(* Logix 5000 project; controller NWGG 1756-L72 rev 35.12; software revision 35.00 *) (continued)

ADD_ON_INSTRUCTION AndcoAnalog   (* revision 1.0 *)
VAR_IN_OUT
   Andco_Values : udt_Andco_Values; {required}
   Andco_Motor_Open : BOOL; {required}
   Anco_Motor_Close : BOOL; {required}
END_VAR
VAR_INPUT
   AnalogValue : DINT; {access Read Only, required}
END_VAR
VAR
   tmr_Web_Watchdog : TIMER := (PRE := 30000); {access None}
   Cal_Open_Gate : BOOL; {access None}
   Cal_Close_Gate : BOOL; {access None}
   Motor_Wind_Down : DINT; {access None}
   Cal_Mid_Point : DINT; {access None}
   Cal_Preact : BOOL; {access None}
   Cal_Finish_Close_Gate : BOOL; {access None}
   tmr_Motor_Wind_Down : TIMER[8] := ([1].PRE := 1000, [2].PRE := 1000); {access None}
   New_Position : DINT; {access None}
   Move_Open : BOOL; {access None}
   Move_Close : BOOL; {access None}
   Adjusted_New_Position : DINT; {access None}
   Cal_Init_Bin_Closed : BOOL; {access None}
   tmrCalCloseGate : TIMER := (PRE := 55000); {access None}
   CurrentPosition : DINT; {access None}
   tmrCalOpenGate : TIMER := (PRE := 55000); {access None}
   CalReturnToPosition : BOOL; {access None}
   CalibratingGate : BOOL; {access None}
   onsStartCal : BOOL; {access None}
   sbCalGateClosed : BOOL; {access None}
   obCalGateClosed : BOOL; {access None}
   sbStartCal : BOOL; {access None}
   obStartCal : BOOL; {access None}
   sbCalGateOpened : BOOL; {access None}
   obCalGateOpened : BOOL; {access None}
END_VAR

ROUTINE Logic   (* ladder *)
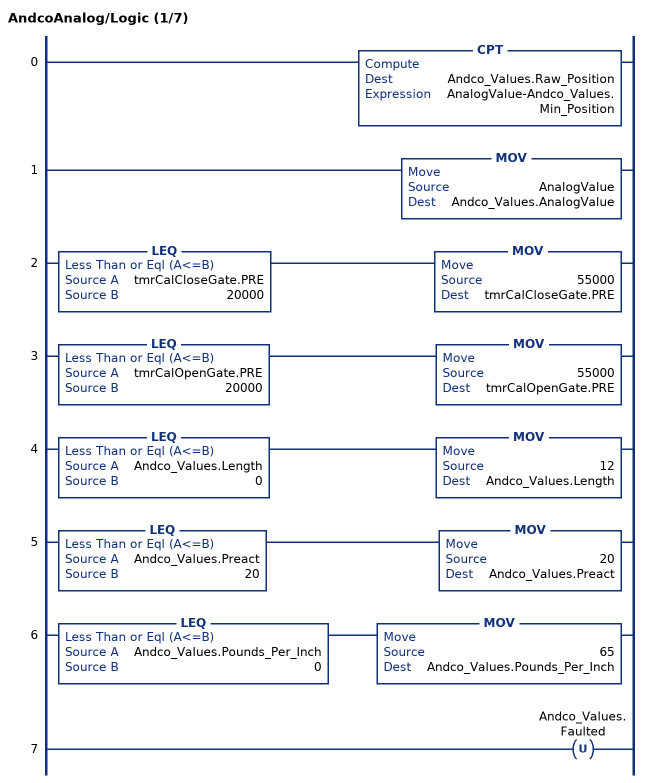
   0: CPT(Andco_Values.Raw_Position,AnalogValue-Andco_Values.Min_Position);
   1: MOV(AnalogValue,Andco_Values.AnalogValue);
   2: LEQ(tmrCalCloseGate.PRE,20000)MOV(55000,tmrCalCloseGate.PRE);
   3: LEQ(tmrCalOpenGate.PRE,20000)MOV(55000,tmrCalOpenGate.PRE);
   4: LEQ(Andco_Values.Length,0)MOV(12,Andco_Values.Length);
   5: LEQ(Andco_Values.Preact,20)MOV(20,Andco_Values.Preact);
   6: LEQ(Andco_Values.Pounds_Per_Inch,0)MOV(65,Andco_Values.Pounds_Per_Inch);
   7: OTU(Andco_Values.Faulted);
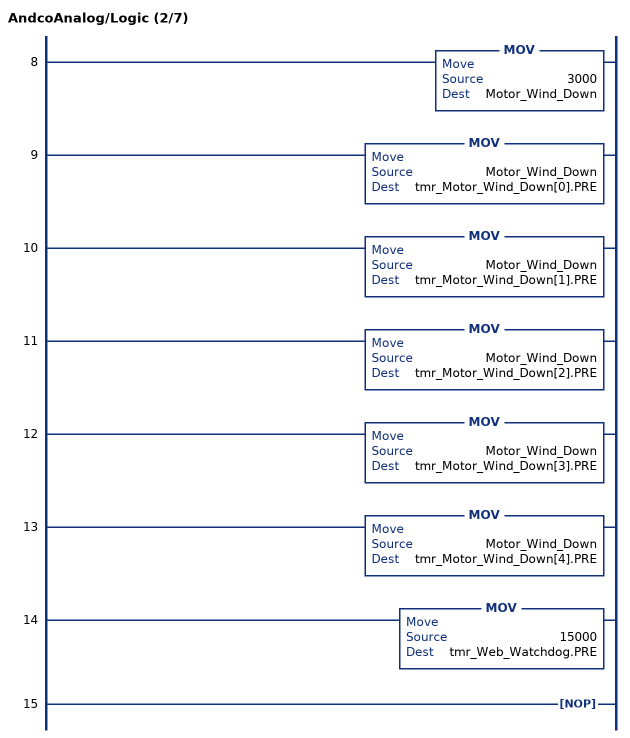
   8: MOV(3000,Motor_Wind_Down);
   9: MOV(Motor_Wind_Down,tmr_Motor_Wind_Down[0].PRE);
   10: MOV(Motor_Wind_Down,tmr_Motor_Wind_Down[1].PRE);
   11: MOV(Motor_Wind_Down,tmr_Motor_Wind_Down[2].PRE);
   12: MOV(Motor_Wind_Down,tmr_Motor_Wind_Down[3].PRE);
   13: MOV(Motor_Wind_Down,tmr_Motor_Wind_Down[4].PRE);
   14: MOV(15000,tmr_Web_Watchdog.PRE);
   15: NOP();
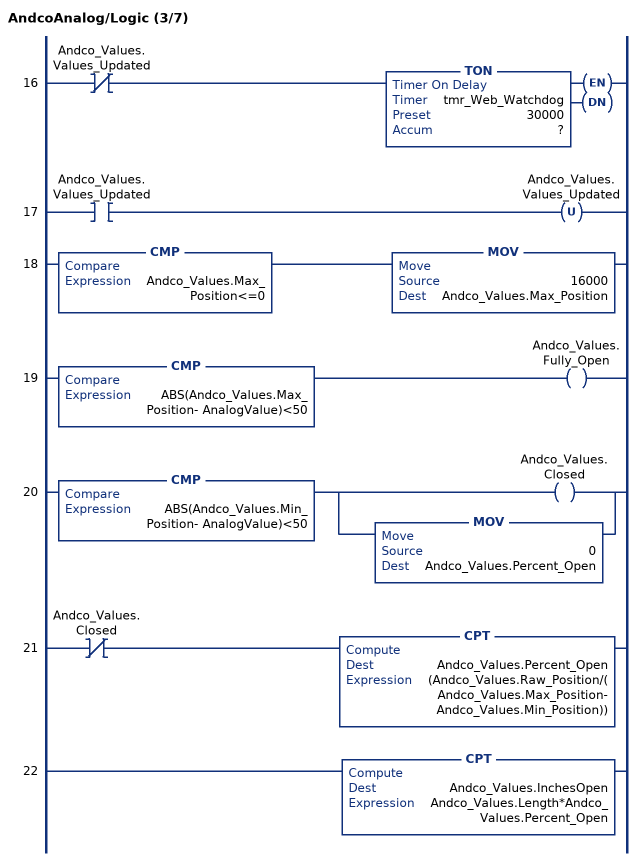
   16: XIO(Andco_Values.Values_Updated)TON(tmr_Web_Watchdog,?,?);
   17: XIC(Andco_Values.Values_Updated)OTU(Andco_Values.Values_Updated);
   18: CMP(Andco_Values.Max_Position<=0)MOV(16000,Andco_Values.Max_Position);
   19: CMP(ABS(Andco_Values.Max_Position- AnalogValue)<50)OTE(Andco_Values.Fully_Open);
   20: CMP(ABS(Andco_Values.Min_Position- AnalogValue)<50)[OTE(Andco_Values.Closed) ,MOV(0,Andco_Values.Percent_Open) ];
   21: XIO(Andco_Values.Closed)CPT(Andco_Values.Percent_Open,(Andco_Values.Raw_Position/(Andco_Values.Max_Position-Andco_Values.Min_Position)));
   22: CPT(Andco_Values.InchesOpen,Andco_Values.Length*Andco_Values.Percent_Open);
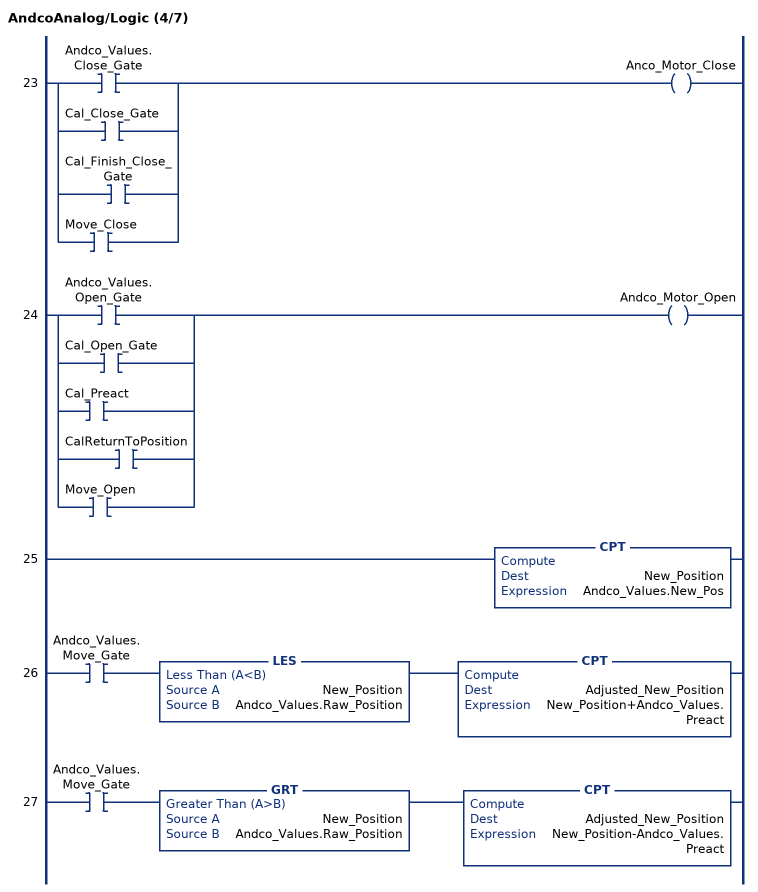
   23: [XIC(Andco_Values.Close_Gate) ,XIC(Cal_Close_Gate) ,XIC(Cal_Finish_Close_Gate) ,XIC(Move_Close) ]OTE(Anco_Motor_Close);
   24: [XIC(Andco_Values.Open_Gate) ,XIC(Cal_Open_Gate) ,XIC(Cal_Preact) ,XIC(CalReturnToPosition) ,XIC(Move_Open) ]OTE(Andco_Motor_Open);
   25: CPT(New_Position,Andco_Values.New_Pos);
   26: XIC(Andco_Values.Move_Gate)LES(New_Position,Andco_Values.Raw_Position)CPT(Adjusted_New_Position,New_Position+Andco_Values.Preact);
   27: XIC(Andco_Values.Move_Gate)GRT(New_Position,Andco_Values.Raw_Position)CPT(Adjusted_New_Position,New_Position-Andco_Values.Preact);
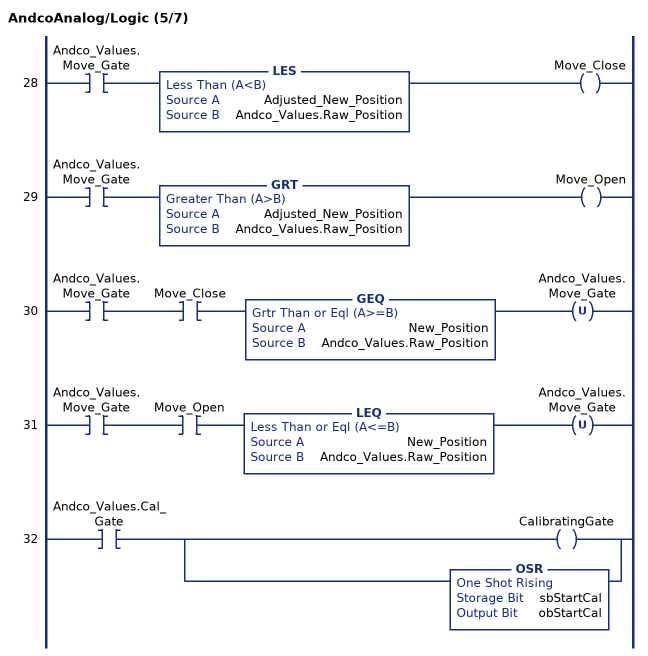
   28: XIC(Andco_Values.Move_Gate)LES(Adjusted_New_Position,Andco_Values.Raw_Position)OTE(Move_Close);
   29: XIC(Andco_Values.Move_Gate)GRT(Adjusted_New_Position,Andco_Values.Raw_Position)OTE(Move_Open);
   30: XIC(Andco_Values.Move_Gate)XIC(Move_Close)GEQ(New_Position,Andco_Values.Raw_Position)OTU(Andco_Values.Move_Gate);
   31: XIC(Andco_Values.Move_Gate)XIC(Move_Open)LEQ(New_Position,Andco_Values.Raw_Position)OTU(Andco_Values.Move_Gate);
   32: XIC(Andco_Values.Cal_Gate)[OTE(CalibratingGate) ,OSR(sbStartCal,obStartCal) ];
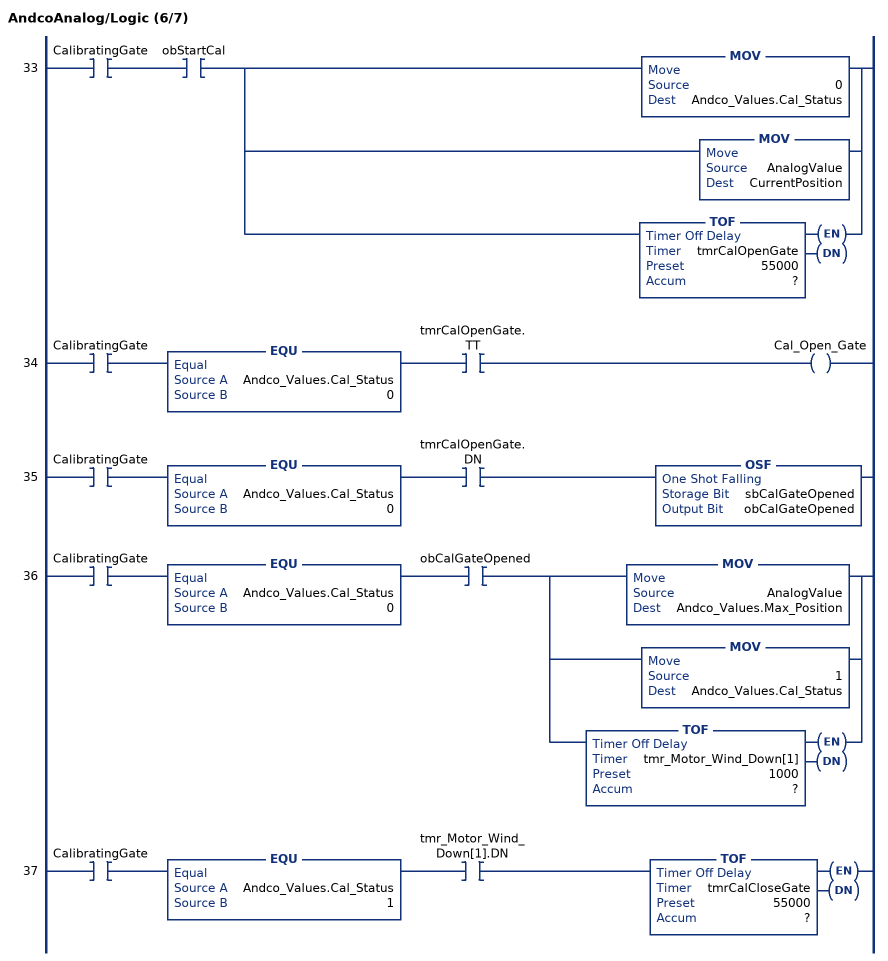
   33: XIC(CalibratingGate)XIC(obStartCal)[MOV(0,Andco_Values.Cal_Status) ,MOV(AnalogValue,CurrentPosition) ,TOF(tmrCalOpenGate,?,?) ];
   34: XIC(CalibratingGate)EQU(Andco_Values.Cal_Status,0)XIC(tmrCalOpenGate.TT)OTE(Cal_Open_Gate);
   35: XIC(CalibratingGate)EQU(Andco_Values.Cal_Status,0)XIC(tmrCalOpenGate.DN)OSF(sbCalGateOpened,obCalGateOpened);
   36: XIC(CalibratingGate)EQU(Andco_Values.Cal_Status,0)XIC(obCalGateOpened)[MOV(AnalogValue,Andco_Values.Max_Position) ,MOV(1,Andco_Values.Cal_Status) ,TOF(tmr_Motor_Wind_Down[1],?,?) ];
   37: XIC(CalibratingGate)EQU(Andco_Values.Cal_Status,1)XIC(tmr_Motor_Wind_Down[1].DN)TOF(tmrCalCloseGate,?,?);
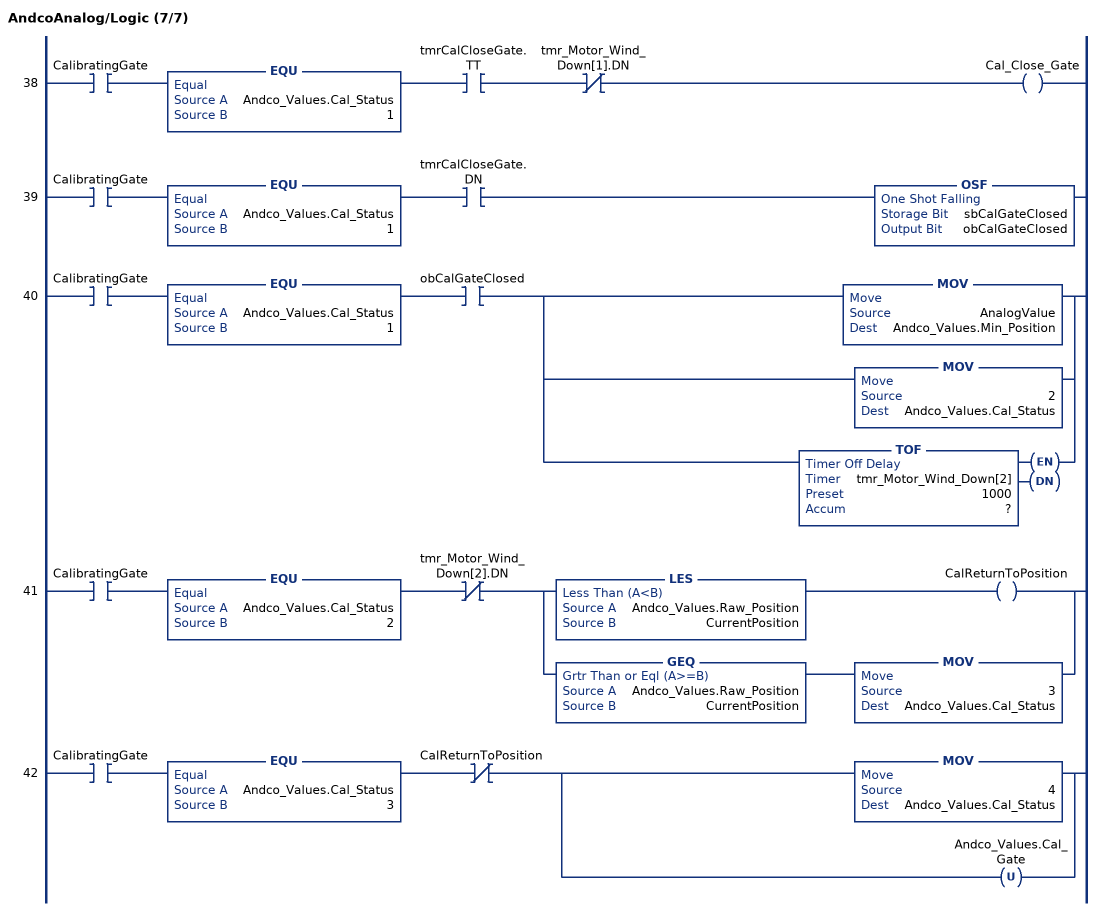
   38: XIC(CalibratingGate)EQU(Andco_Values.Cal_Status,1)XIC(tmrCalCloseGate.TT)XIO(tmr_Motor_Wind_Down[1].DN)OTE(Cal_Close_Gate);
   39: XIC(CalibratingGate)EQU(Andco_Values.Cal_Status,1)XIC(tmrCalCloseGate.DN)OSF(sbCalGateClosed,obCalGateClosed);
   40: XIC(CalibratingGate)EQU(Andco_Values.Cal_Status,1)XIC(obCalGateClosed)[MOV(AnalogValue,Andco_Values.Min_Position) ,MOV(2,Andco_Values.Cal_Status) ,TOF(tmr_Motor_Wind_Down[2],?,?) ];
   41: XIC(CalibratingGate)EQU(Andco_Values.Cal_Status,2)XIO(tmr_Motor_Wind_Down[2].DN)[LES(Andco_Values.Raw_Position,CurrentPosition) OTE(CalReturnToPosition) ,GEQ(Andco_Values.Raw_Position,CurrentPosition) MOV(3,Andco_Values.Cal_Status) ];
   42: XIC(CalibratingGate)EQU(Andco_Values.Cal_Status,3)XIO(CalReturnToPosition)[MOV(4,Andco_Values.Cal_Status) ,OTU(Andco_Values.Cal_Gate) ];
END_ROUTINE
END_ADD_ON_INSTRUCTION

ADD_ON_INSTRUCTION HOUR_METER   (* revision 1.0 *)
VAR_INPUT
   MOTOR_RUNNING_INPUT_1 : BOOL; {required}
END_VAR
VAR_OUTPUT
   HR_METER_DISPLAY : DINT; {visible}
END_VAR
VAR_INPUT
   NEXT_SCHDL_MAINTENANCE : DINT; {visible}
END_VAR
VAR_OUTPUT
   MAINTENANCE_ALARM : BOOL; {visible}
END_VAR
VAR
   COUNTER : COUNTER := (PRE := 99999999); {access None}
   TIMER : TIMER := (PRE := 3600000); {access None}
END_VAR

ROUTINE Logic   (* ladder *)
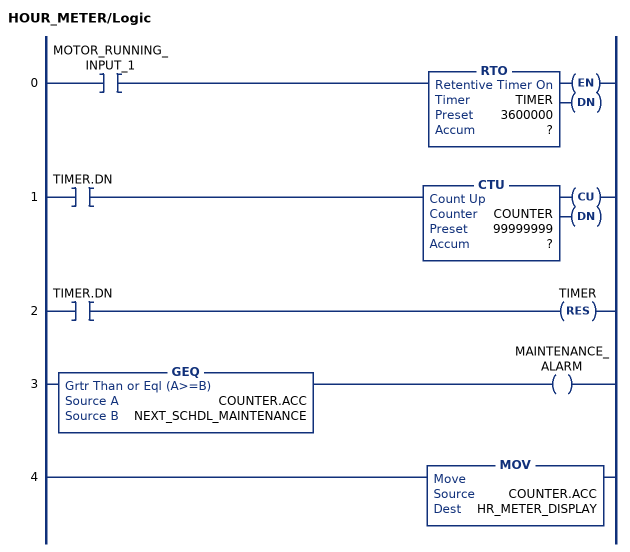
   0: XIC(MOTOR_RUNNING_INPUT_1)RTO(TIMER,?,?);
   1: XIC(TIMER.DN)CTU(COUNTER,?,?);
   2: XIC(TIMER.DN)RES(TIMER);
   3: GEQ(COUNTER.ACC,NEXT_SCHDL_MAINTENANCE)OTE(MAINTENANCE_ALARM);
   4: MOV(COUNTER.ACC,HR_METER_DISPLAY);
END_ROUTINE
END_ADD_ON_INSTRUCTION

ADD_ON_INSTRUCTION Loadout_Bin_Control   (* revision 1.0 *)
VAR_IN_OUT
   Bin : udt_Loadout_Bin; {required}
   Open_Air_Gate : BOOL; {required}
END_VAR
VAR_INPUT
   Bin_Open_Treat_Pause : BOOL; {required}
   Bin_Open_Clean_Pause : BOOL; {required}
END_VAR
VAR_IN_OUT
   TMR_Max_Treat_Delay : TIMER; {required}
   TMR_Max_Clean_Delay : TIMER; {required}
   Air_Gate_Open_Input : BOOL; {required}
   Auger_Relay : BOOL; {required}
END_VAR
VAR_INPUT
   Use_Auger_Relay : BOOL; {required}
   Use_Bindicator : BOOL; {access None, required}
END_VAR
VAR_IN_OUT
   Bindicator_Input : BOOL; {required}
   ALM_Air_Gate_Failed : ALARM_DIGITAL; {required}
END_VAR
VAR_INPUT
   Bin_Open_Transfer_Pause : BOOL; {required}
END_VAR
VAR_IN_OUT
   Clean_Batch_Status : DINT; {required}
   Treat_Batch_Status : DINT; {required}
   Transfer_Batch_Status : DINT; {required}
   Andco_Motor_Open : BOOL; {required}
   Andco_Motor_Close : BOOL; {required}
   Required_Belt : BOOL; {required}
   Manual_Mode : BOOL; {required}
END_VAR
VAR_INPUT
   RawAnalogTag : DINT; {access Read Only, required}
END_VAR
VAR
   Auto_Open_Air_Gate_Ready : BOOL; {access None}
   Air_Gate_Open_Cal : BOOL; {access None}
   TMR_Air_Gate_Fail : TIMER := (PRE := 4000); {access None}
   ALM_Air_Gate_Failed_Ack : BOOL; {access None}
   Air_Gate_Open_Clean : BOOL; {access None}
   Air_Gate_Open_Treat : BOOL; {access None}
   Air_Gate_Open_Transfer : BOOL; {access None}
   Andco : Andco; {access None}
   Open_Treat_Air_Gate : BOOL; {access None}
   Open_Treat_Air_Gate_Ready : BOOL; {access None}
   AndcoAnalog : AndcoAnalog; {access None}
END_VAR

ROUTINE Logic   (* ladder *)
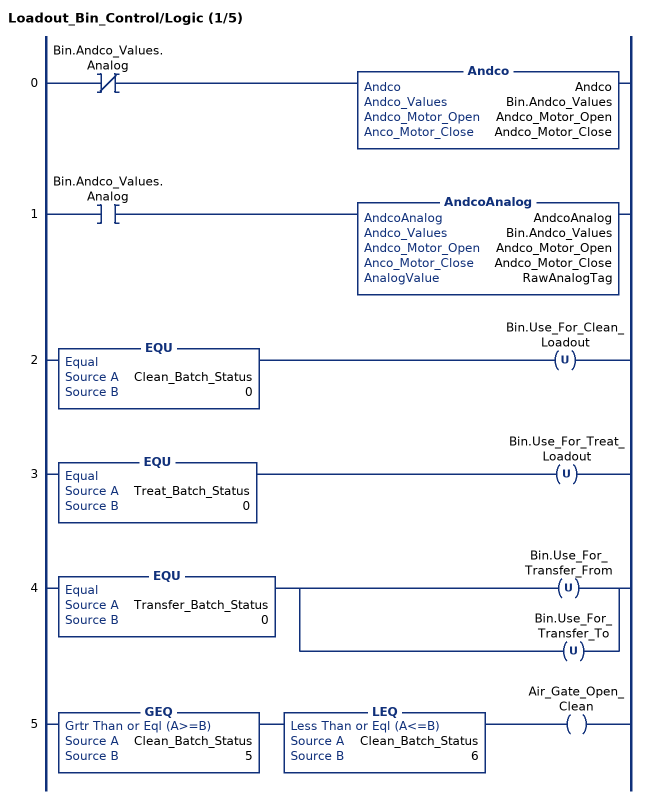
   0: XIO(Bin.Andco_Values.Analog)Andco(Andco,Bin.Andco_Values,Andco_Motor_Open,Andco_Motor_Close);
   1: XIC(Bin.Andco_Values.Analog)AndcoAnalog(AndcoAnalog,Bin.Andco_Values,Andco_Motor_Open,Andco_Motor_Close,RawAnalogTag);
   2: EQU(Clean_Batch_Status,0)OTU(Bin.Use_For_Clean_Loadout);
   3: EQU(Treat_Batch_Status,0)OTU(Bin.Use_For_Treat_Loadout);
   4: EQU(Transfer_Batch_Status,0)[OTU(Bin.Use_For_Transfer_From) ,OTU(Bin.Use_For_Transfer_To) ];
   5: GEQ(Clean_Batch_Status,5)LEQ(Clean_Batch_Status,6)OTE(Air_Gate_Open_Clean);
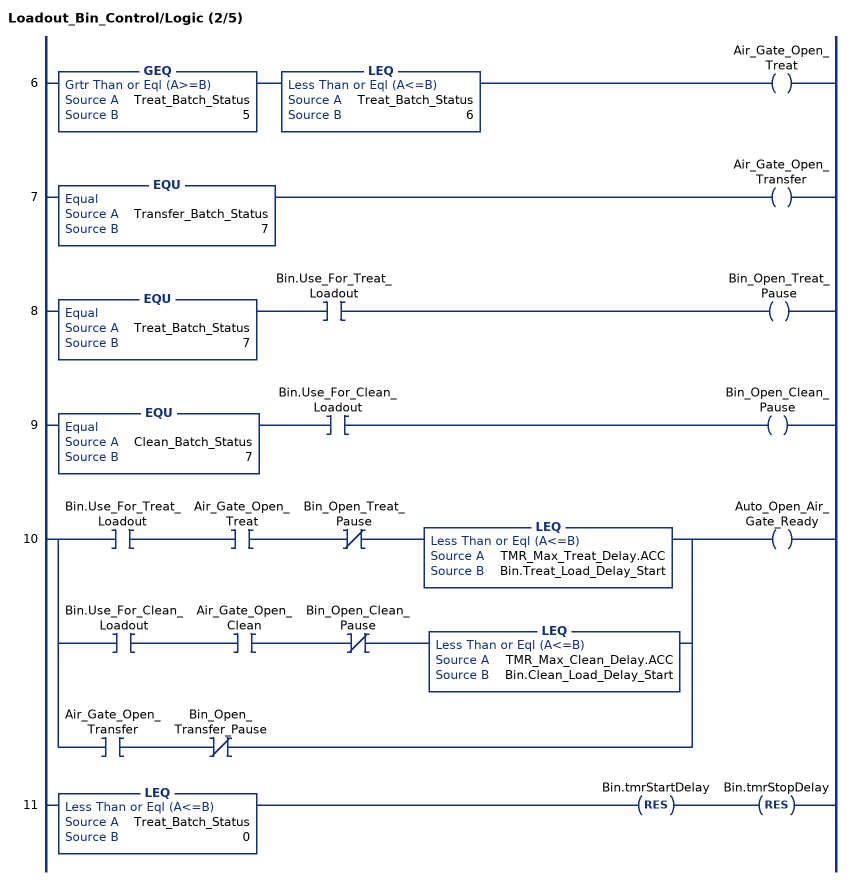
   6: GEQ(Treat_Batch_Status,5)LEQ(Treat_Batch_Status,6)OTE(Air_Gate_Open_Treat);
   7: EQU(Transfer_Batch_Status,7)OTE(Air_Gate_Open_Transfer);
   8: EQU(Treat_Batch_Status,7)XIC(Bin.Use_For_Treat_Loadout)OTE(Bin_Open_Treat_Pause);
   9: EQU(Clean_Batch_Status,7)XIC(Bin.Use_For_Clean_Loadout)OTE(Bin_Open_Clean_Pause);
   10: [XIC(Bin.Use_For_Treat_Loadout) XIC(Air_Gate_Open_Treat) XIO(Bin_Open_Treat_Pause) LEQ(TMR_Max_Treat_Delay.ACC,Bin.Treat_Load_Delay_Start) ,XIC(Bin.Use_For_Clean_Loadout) XIC(Air_Gate_Open_Clean) XIO(Bin_Open_Clean_Pause) LEQ(TMR_Max_Clean_Delay.ACC,Bin.Clean_Load_Delay_Start) ,XIC(Air_Gate_Open_Transfer) XIO(Bin_Open_Transfer_Pause) ]OTE(Auto_Open_Air_Gate_Ready);
   11: LEQ(Treat_Batch_Status,0)RES(Bin.tmrStartDelay)RES(Bin.tmrStopDelay);
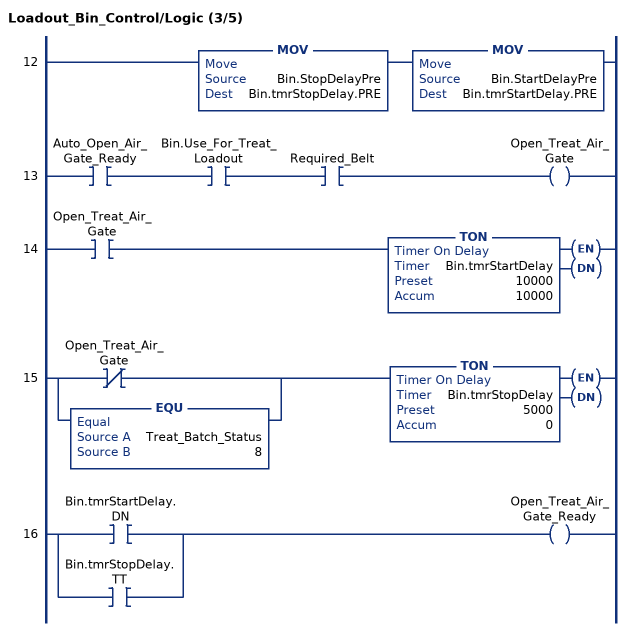
   12: MOV(Bin.StopDelayPre,Bin.tmrStopDelay.PRE)MOV(Bin.StartDelayPre,Bin.tmrStartDelay.PRE);
   13: XIC(Auto_Open_Air_Gate_Ready)XIC(Bin.Use_For_Treat_Loadout)XIC(Required_Belt)OTE(Open_Treat_Air_Gate);
   14: XIC(Open_Treat_Air_Gate)TON(Bin.tmrStartDelay,10000,10000);
   15: [XIO(Open_Treat_Air_Gate) ,EQU(Treat_Batch_Status,8) ]TON(Bin.tmrStopDelay,5000,0);
   16: [XIC(Bin.tmrStartDelay.DN) ,XIC(Bin.tmrStopDelay.TT) ]OTE(Open_Treat_Air_Gate_Ready);
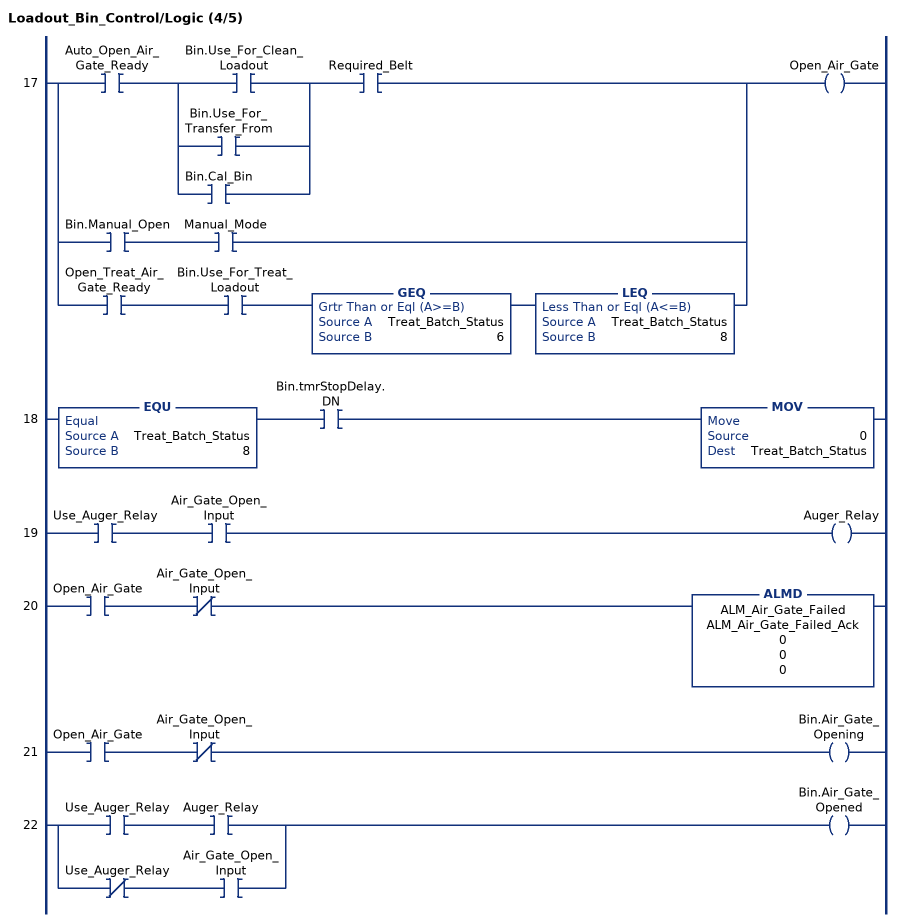
   17: [XIC(Auto_Open_Air_Gate_Ready) [XIC(Bin.Use_For_Clean_Loadout) ,XIC(Bin.Use_For_Transfer_From) ,XIC(Bin.Cal_Bin) ] XIC(Required_Belt) ,XIC(Bin.Manual_Open) XIC(Manual_Mode) ,XIC(Open_Treat_Air_Gate_Ready) XIC(Bin.Use_For_Treat_Loadout) GEQ(Treat_Batch_Status,6) LEQ(Treat_Batch_Status,8) ]OTE(Open_Air_Gate);
   18: EQU(Treat_Batch_Status,8)XIC(Bin.tmrStopDelay.DN)MOV(0,Treat_Batch_Status);
   19: XIC(Use_Auger_Relay)XIC(Air_Gate_Open_Input)OTE(Auger_Relay);
   20: XIC(Open_Air_Gate)XIO(Air_Gate_Open_Input)ALMD(ALM_Air_Gate_Failed,ALM_Air_Gate_Failed_Ack,0,0,0);
   21: XIC(Open_Air_Gate)XIO(Air_Gate_Open_Input)OTE(Bin.Air_Gate_Opening);
   22: [XIC(Use_Auger_Relay) XIC(Auger_Relay) ,XIO(Use_Auger_Relay) XIC(Air_Gate_Open_Input) ]OTE(Bin.Air_Gate_Opened);
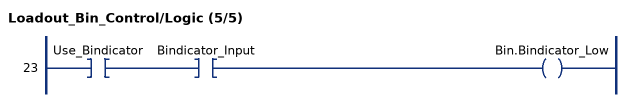
   23: XIC(Use_Bindicator)XIC(Bindicator_Input)OTE(Bin.Bindicator_Low);
END_ROUTINE
END_ADD_ON_INSTRUCTION
